// TIA Portal project "Test_PID_Level" (V15.1)

(* hardware
DEVICE "S71500/ET200MP station_1"  S7-1500 station
   slot 0: "Telaio di montaggio_0"  Rack  6ES7 590-1***0-0AA0
   slot 1: "PLC_1"  CPU 1515-2 PN  6ES7 515-2AM01-0AB0  V2.6
      slot 3: "Display CPU_1"  6ES7591-1BA00-0AA0
DEVICE "HMI_1"  TP2200 Comfort
   slot 0: "HMI_1"  TP2200 Comfort  6AV2 124-0XC02-0AX1  15.1.0.0
   slot 1: "HMI_RT_1"  TP2200 Comfort  6AV2 124-0XC02-0AX1  15.1.0.0
   slot 5: "HMI_1.IE_CP_1"  PROFINET Interface  15.0.1.0
      slot 1: "Interfaccia_1 PROFINET"  PROFINET Interface
         slot 1: "Porta_1"  Port
         slot 2: "Porta_2"  Port
   slot 6: "HMI_1.IE_CP_2"  PROFINET Interface  15.0.1.0
      slot 1: "PROFINET Interface_GBit"  PROFINET Interface
         slot 1: "Porta_1"  Port
   slot 7: "HMI_1.MPI/DP_CP_1"  MPI/DP Interface  15.0.1.0
*)

// ===== PLC "PLC_1"  CPU 1515-2 PN =====

TYPE "s_PID"
   STRUCT
      i_Set_Point : Real;   // Set point value
      i_Feedback : Real;   // Feedback value process
      i_Kp : Real;   // K Proportional gain
      i_Ki : Real;   // K Integral gain
      i_Kd : Real;   // K Derivative gain
      i_Max_Analog : Real;   // Maximum value for analog output
      i_Duty_Cycle : Real;   // Maximum time cycle for PWM digital output (milliseconds)
      i_Scan_Time : Real;   // Scanning time of the plc
      i_Time_Sample : Real;   // Time sample in OB35
      i_Enable_PWM : Bool;   // Enable PWM digital P.I.D.
      i_Reset : Bool;   // Reset regulator
      i_Enable_I : Bool;   // Enable Integral component
      o_Analog_Reg : Real;   // Output analog regulation
      o_Duty_Cycle_Perc : Real;   // Duty cycle On percentage
      o_Wave_On_PWM : Bool;   // Output high wave On of digital PWM
      o_Wave_Off_PWM : Bool;   // Output low wave On of digital PWM
   END_STRUCT;
END_TYPE

DATA_BLOCK "f_PID_DB"   // DB80
{ S7_Optimized_Access := 'TRUE' }
VERSION : 0.1
// stored: InstanceOfName f_PID
"f_PID"
BEGIN
END_DATA_BLOCK

DATA_BLOCK "DB_PID"   // DB82
{ S7_Optimized_Access := 'TRUE' }
VERSION : 0.1
   VAR RETAIN
      Data : "s_PID";   // Valve 1
   END_VAR
   VAR
      Scan_Time_LR : LReal;
      Mem_Scan_Time : LReal;
      Scan_Time_R : Real;
      FB_Int : Int;
      Derivative_ON : Bool;
      Enable_I : Bool;
   END_VAR
BEGIN
END_DATA_BLOCK

DATA_BLOCK "DB_Tank"   // DB83
{ S7_Optimized_Access := 'TRUE' }
VERSION : 0.1
   VAR
      V1_On : Bool;
      V2_On : Bool;
      V3_On : Bool;
      V4_On : Bool;
      V1_Max : Real;   // Liters per second V1, input
      V2_SP : Real;   // Set point Liters per second
      V3_SP : Real;   // Set point Liters per second
      V4_SP : Real;   // Set point Liters per second
      Water : Real;   // Liters
      Tank_Max : Real := 3000.0;
      V1_In : Real;   // Liters in input
      V2_Out : Real;   // Liters in output
      V3_Out : Real;   // Liters in output
      V4_Out : Real;   // Liters in output
      FB_V1 : Real;
   END_VAR
BEGIN
END_DATA_BLOCK

FUNCTION_BLOCK "f_PID"   // FB80, SCL
{ S7_Optimized_Access := 'TRUE' }
VERSION : 0.1
   VAR_INPUT
      Set_Point : Real;   // Set point value
      Feedback : Real;   // Feedback value process
      Kp : Real;   // K Proportional gain
      Ki : Real;   // K Integral gain
      Kd : Real;   // K Derivative gain
      Max_Analog : Real;   // Maximum value for analog output
      Duty_Cycle : Real;   // Maximum time cycle for PWM digital output (milliseconds)
      Scan_Time : Real;   // Scanning time of the plc
      Time_Sample : Real;   // Time sample in OB35
      Enable_PWM : Bool;   // Enable PWM digital P.I.D.
      Reset : Bool;   // Reset regulator
      Enable_I : Bool;
   END_VAR
   VAR_OUTPUT
      Analog_Reg : Real;   // Output analog regulation
      Duty_Cycle_Perc : Real;   // Duty cycle On percentage
      Wave_On_PWM : Bool;   // Output high wave On of digital PWM
      Wave_Off_PWM : Bool;   // Output low wave On of digital PWM
      Derivative_ON : Bool;
   END_VAR
   VAR
      Error : Real;   // Error for each scan
      I_Ist : Real;   // Istant integral
      I : Real;   // Integral component
      D : Real;   // Derivative component
      P : Real;   // Proportional component
      Last_Error : Real;   // Error of previous scan
      Accu_Timer : Real;   // Timer Accumulator for the duty cycle PWM
      Thr_Wave_On : Real;   // Threshold for the wave ON
      Thr_Wave_Off : Real;   // Threshold for the wave OFF
      Wave_On : Bool;   // Wave On
      Wave_Off : Bool;   // Wave Off
   END_VAR
BEGIN
   // P.I.D. Regulator. Written By Ing. Walter Porcellini Milan (Italy) the 15/09/2021
   // I revisited and modified the algorithm I wrote in June 2009
   // This project and its algorithm are intended as a didactic demonstration
   // I decline from any responsibility for damage to things and / or people.

   #Error := #Set_Point - #Feedback;

   #P := #Error * #Kp * 1.0;

   IF #P > #Max_Analog THEN

       #P := #Max_Analog;
   END_IF;

   IF #P < (#Max_Analog * -1.0) THEN

       #P := #Max_Analog * -1.0;
   END_IF;

   IF #Enable_I = true THEN
       #I_Ist := #Error * #Ki * 1.0;
       #I := #I + #I_Ist;

   ELSE
       #I_Ist := 0.0;
       #I := 0.0;
   END_IF;

   #I := #I + #I_Ist;

   IF #I <= 0.0 THEN
      #I := 0.0;
   END_IF;

   IF #I >= #Max_Analog * 0.8 THEN
       #I := #Max_Analog * 0.8;
   END_IF;

   IF #Time_Sample > 0.0 THEN
       #D := (#Kd * 1.0*(#Error - #Last_Error)) / #Time_Sample;
   END_IF;

   #Last_Error := #Error;

   #Analog_Reg := #P + #I + #D;

   #Derivative_ON := #D <> 0.0;

   IF #Reset THEN

       #P := 0.0;
       #I := 0.0;
       #I_Ist := 0.0;
       #D := 0.0;
       #Analog_Reg := 0.0;
       #Wave_On := false;
       #Wave_Off := false;
       #Accu_Timer := 0.0;
       #Last_Error := 0.0;

   END_IF;

   IF #Analog_Reg >= #Max_Analog THEN
       #Analog_Reg := #Max_Analog;
   END_IF;

   IF #Analog_Reg <= 0.0 THEN
       #Analog_Reg:=0.0;
   END_IF;


   IF #Enable_PWM = true THEN
       #Thr_Wave_On := (#Duty_Cycle / #Max_Analog) * #Analog_Reg;

       #Thr_Wave_Off := #Max_Analog - #Thr_Wave_On;


       IF #Accu_Timer = 0.0 AND #Enable_PWM = TRUE THEN

           #Wave_On := true;
           #Wave_Off := false;

       END_IF;

       IF #Wave_On = true THEN

           #Accu_Timer := #Accu_Timer + #Time_Sample;
           #Duty_Cycle_Perc := (#Thr_Wave_On / #Duty_Cycle) * 100.0;

           IF #Accu_Timer >= #Thr_Wave_On THEN

               #Wave_On := false;
               #Wave_Off := true;

           END_IF;

       END_IF;


       IF #Wave_Off = true THEN

           #Accu_Timer := #Accu_Timer + #Time_Sample;

           IF #Accu_Timer >= #Duty_Cycle THEN

               #Wave_Off := false;
               #Accu_Timer := 0.0;

           END_IF;

       END_IF;



       #Wave_On_PWM := #Wave_On AND #Thr_Wave_On >= 1000.0;
       #Wave_Off_PWM := #Wave_Off;

   ELSE
       #Wave_On_PWM := false;
       #Wave_Off_PWM := false;
       #Accu_Timer := 0.0;
       #Duty_Cycle_Perc := 0.0;
   END_IF;
END_FUNCTION_BLOCK

FUNCTION "1_Temperature" : Void   // FC100, SCL
{ S7_Optimized_Access := 'TRUE' }
VERSION : 0.1
BEGIN
   // "DB_PID".V1.i_Feedback := INT_TO_REAL("DB_PID".FB_Int);

   "DB_PID".Data.i_Feedback := "DB_PID".Data.i_Feedback + ("DB_PID".Data.o_Analog_Reg * 0.000000024);
   "DB_PID".Data.i_Feedback := "DB_PID".Data.i_Feedback - 0.00008;

   IF "DB_PID".Data.i_Feedback < 20.0 OR "DB_PID".Data.i_Reset = true THEN

       "DB_PID".Data.i_Feedback := 20.0;
   END_IF;


   IF "DB_PID".Data.i_Feedback > 150.0 THEN

       "DB_PID".Data.i_Feedback := 150.0;
   END_IF;
END_FUNCTION

FUNCTION "2_Tank Level" : Void   // FC101, SCL
{ S7_Optimized_Access := 'TRUE' }
VERSION : 0.1
   VAR_TEMP
      Stop_Integral : Bool;
   END_VAR
BEGIN

   IF "DB_Tank".V2_SP > 30.0 THEN

       "DB_Tank".V2_SP := 30.0;

   END_IF;

   IF "DB_Tank".V2_SP < 0.0 THEN

       "DB_Tank".V2_SP := 0.0;

   END_IF;

   IF "DB_Tank".V3_SP > 30.0 THEN

       "DB_Tank".V3_SP := 30.0;

   END_IF;

   IF "DB_Tank".V3_SP < 0.0 THEN

       "DB_Tank".V3_SP := 0.0;

   END_IF;

   IF "DB_Tank".V4_SP > 30.0 THEN

       "DB_Tank".V4_SP := 30.0;

   END_IF;

   IF "DB_Tank".V4_SP < 0.0 THEN

       "DB_Tank".V4_SP := 0.0;

   END_IF;

   "DB_Tank".V2_Out := ("DB_Tank".V2_SP * "DB_PID".Scan_Time_R);
   "DB_Tank".V3_Out := ("DB_Tank".V3_SP * "DB_PID".Scan_Time_R);
   "DB_Tank".V4_Out := ("DB_Tank".V4_SP * "DB_PID".Scan_Time_R);

   IF "DB_Tank".V2_On = true THEN
       "DB_Tank".Water := "DB_Tank".Water - "DB_Tank".V2_Out;

   END_IF;

   IF "DB_Tank".V3_On = true THEN
       "DB_Tank".Water := "DB_Tank".Water - "DB_Tank".V3_Out;

   END_IF;

   IF "DB_Tank".V4_On = true THEN
       "DB_Tank".Water := "DB_Tank".Water - "DB_Tank".V4_Out;

   END_IF;

   "DB_Tank".V1_Max := 100.0;
   "DB_Tank".V1_In := ("DB_Tank".V1_Max / "DB_PID".Data.i_Max_Analog) * "DB_PID".Data.o_Analog_Reg * "DB_PID".Scan_Time_R ;
   "DB_Tank".FB_V1 := "DB_Tank".V1_In * 1000.0;

   "DB_Tank".Water := "DB_Tank".Water + "DB_Tank".V1_In;

   IF "DB_Tank".Water < 0.0 OR "DB_PID".Data.i_Reset=true THEN

       "DB_Tank".Water := 0;
   END_IF;

   "DB_Tank".V1_On := "DB_PID".Data.o_Analog_Reg > 0.0;
   "DB_PID".Data.i_Feedback := "DB_Tank".Water;
   "DB_PID".FB_Int := REAL_TO_INT("DB_Tank".Water);

   #Stop_Integral := "DB_Tank".V2_On = false
   AND "DB_Tank".V3_On = false
   AND "DB_Tank".V4_On = false;

   "DB_PID".Enable_I := NOT #Stop_Integral;
END_FUNCTION

ORGANIZATION_BLOCK "Main"   // OB1, LAD, ProgramCycle
TITLE = "Main Program Sweep (Cycle)"
{ S7_Optimized_Access := 'TRUE' }
VERSION : 0.1
   VAR_INPUT
      Initial_Call : Bool;   // Initial call of this OB
      Remanence : Bool;   // =True, if remanent data are available
   END_VAR
BEGIN

REGION Network 1
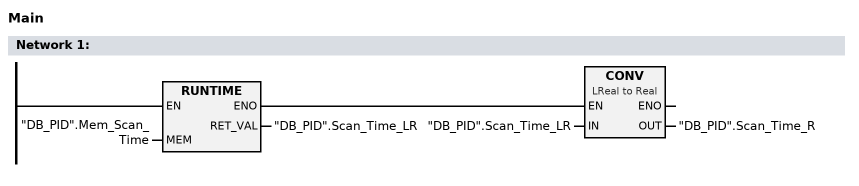
   // no SCL statement known for Runtime: written as a call
   // ENO of a box is taken as its EN; it also drops when the box reports an error
   "DB_PID".Scan_Time_LR := Runtime(mem := "DB_PID".Mem_Scan_Time);
   "DB_PID".Scan_Time_R := LREAL_TO_REAL("DB_PID".Scan_Time_LR);
END_REGION

REGION Network 2 (SCL)
   "DB_PID".Data.i_Max_Analog := 16384;
   "DB_PID".Data.i_Duty_Cycle := 10000;
   "DB_PID".Data.i_Scan_Time := "DB_PID".Scan_Time_R;
   "DB_PID".Data.i_Time_Sample := 10;

   //"1_Temperature"();
   "2_Tank Level"();
END_REGION
END_ORGANIZATION_BLOCK

ORGANIZATION_BLOCK "Cyclic interrupt"   // OB30, LAD, CyclicInterrupt
{ S7_Optimized_Access := 'TRUE' }
VERSION : 0.1
   VAR_INPUT
      Initial_Call : Bool;   // Initial call of this OB
      Event_Count : Int;   // Events discarded
   END_VAR
BEGIN

REGION Network 1
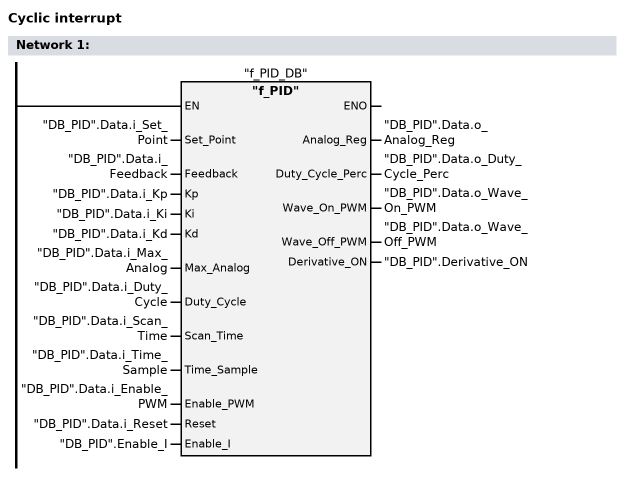
   RUNG wire#powerrail
      "f_PID_DB"(Set_Point := "DB_PID".Data.i_Set_Point, Feedback := "DB_PID".Data.i_Feedback, Kp := "DB_PID".Data.i_Kp, Ki := "DB_PID".Data.i_Ki, Kd := "DB_PID".Data.i_Kd, Max_Analog := "DB_PID".Data.i_Max_Analog, Duty_Cycle := "DB_PID".Data.i_Duty_Cycle, Scan_Time := "DB_PID".Data.i_Scan_Time, Time_Sample := "DB_PID".Data.i_Time_Sample, Enable_PWM := "DB_PID".Data.i_Enable_PWM, Reset := "DB_PID".Data.i_Reset, Enable_I := "DB_PID".Enable_I, Analog_Reg => "DB_PID".Data.o_Analog_Reg, Duty_Cycle_Perc => "DB_PID".Data.o_Duty_Cycle_Perc, Wave_On_PWM => "DB_PID".Data.o_Wave_On_PWM, Wave_Off_PWM => "DB_PID".Data.o_Wave_Off_PWM, Derivative_ON => "DB_PID".Derivative_ON)
   END_RUNG
   // the same network as SCL:
   "f_PID_DB"(Set_Point := "DB_PID".Data.i_Set_Point,   // "f_PID"
              Feedback := "DB_PID".Data.i_Feedback,
              Kp := "DB_PID".Data.i_Kp,
              Ki := "DB_PID".Data.i_Ki,
              Kd := "DB_PID".Data.i_Kd,
              Max_Analog := "DB_PID".Data.i_Max_Analog,
              Duty_Cycle := "DB_PID".Data.i_Duty_Cycle,
              Scan_Time := "DB_PID".Data.i_Scan_Time,
              Time_Sample := "DB_PID".Data.i_Time_Sample,
              Enable_PWM := "DB_PID".Data.i_Enable_PWM,
              Reset := "DB_PID".Data.i_Reset,
              Enable_I := "DB_PID".Enable_I,
              Analog_Reg => "DB_PID".Data.o_Analog_Reg,
              Duty_Cycle_Perc => "DB_PID".Data.o_Duty_Cycle_Perc,
              Wave_On_PWM => "DB_PID".Data.o_Wave_On_PWM,
              Wave_Off_PWM => "DB_PID".Data.o_Wave_Off_PWM,
              Derivative_ON => "DB_PID".Derivative_ON);
END_REGION
END_ORGANIZATION_BLOCK

(* ===== HMI "HMI_RT_1" =====
system functions are stored by id; their names below are inferred from use
connection "HMI_Collegamento_1": ETHERNET, S7_1500_OMS

HMI tags "Tabella delle variabili standard"
   "Variabile_Numero di pagina" : UInt, internal
   "DB_PID_V1_i_Set_Point" : Real = PLC DB_PID.Data.i_Set_Point, 1 s
   "DB_PID_V1_i_Kp" : Real = PLC DB_PID.Data.i_Kp, 1 s
   "DB_PID_V1_i_Feedback" : Real = PLC DB_PID.Data.i_Feedback, 1 s
   "DB_PID_V1_i_Ki" : Real = PLC DB_PID.Data.i_Ki, 1 s
   "DB_PID_V1_i_Kd" : Real = PLC DB_PID.Data.i_Kd, 1 s
   "DB_PID_V1_i_Enable_PWM" : Bool = PLC DB_PID.Data.i_Enable_PWM, 1 s
   "DB_PID_V1_i_Reset" : Bool = PLC DB_PID.Data.i_Reset, 1 s
   "DB_PID_V1_o_Analog_Reg" : Real = PLC DB_PID.Data.o_Analog_Reg, 1 s
   "DB_PID_V1_o_Duty_Cycle_Perc" : Real = PLC DB_PID.Data.o_Duty_Cycle_Perc, 1 s
   "DB_PID_V1_o_Wave_On_PWM" : Bool = PLC DB_PID.Data.o_Wave_On_PWM, 1 s
   "DB_PID_V1_o_Wave_Off_PWM" : Bool = PLC DB_PID.Data.o_Wave_Off_PWM, 1 s
   "DB_PID_FB_Int" : Int = PLC DB_PID.FB_Int, 1 s
   "DB_PID_Derivative_ON" : Bool = PLC DB_PID.Derivative_ON, 1 s
   "DB_Tank_V1_On" : Bool = PLC DB_Tank.V1_On, 1 s
   "DB_Tank_V2_On" : Bool = PLC DB_Tank.V2_On, 1 s
   "DB_Tank_V3_On" : Bool = PLC DB_Tank.V3_On, 1 s
   "DB_Tank_V4_On" : Bool = PLC DB_Tank.V4_On, 1 s
   "DB_Tank_V2_SP" : Real = PLC DB_Tank.V2_SP, 1 s
   "DB_Tank_V3_SP" : Real = PLC DB_Tank.V3_SP, 1 s
   "DB_Tank_V4_SP" : Real = PLC DB_Tank.V4_SP, 1 s
   "f_PID_DB_P" : Real = PLC f_PID_DB.P, 1 s
   "f_PID_DB_I" : Real = PLC f_PID_DB.I, 1 s
   "f_PID_DB_D" : Real = PLC f_PID_DB.D, 1 s
   "DB_Tank_V1_In" : Real = PLC DB_Tank.V1_In, 1 s
   "DB_Tank_FB_V1" : Real = PLC DB_Tank.FB_V1, 1 s

text list "Elenco testi_Nome della pagina": 1 'Pagina base'

screen "Pagina base" 1920x1017, template "Modello_1"
   on GenerateScreen: SetTag("Variabile_Numero di pagina", 1)
   TextField "Casella di testo_1" at 9,24 size 98x25; Text 'Set Point'
   IOField "Campo I/O_1" at 114,21 size 96x32; FormatPattern 9999.9
      ProcessValue <- "DB_PID_V1_i_Set_Point"
   TextField "Casella di testo_2" at 9,68 size 30x25; Text 'Kp'
   IOField "Campo I/O_2" at 114,64 size 96x32; FormatPattern 9999.9
      ProcessValue <- "DB_PID_V1_i_Kp"
   TextField "Casella di testo_3" at 9,111 size 24x25; Text 'Ki'
   IOField "Campo I/O_3" at 114,108 size 96x32; FormatPattern 9999.9
      ProcessValue <- "DB_PID_V1_i_Ki"
   TextField "Casella di testo_4" at 9,155 size 30x25; Text 'Kd'
   IOField "Campo I/O_4" at 114,151 size 96x32; FormatPattern 9999.9
      ProcessValue <- "DB_PID_V1_i_Kd"
   TextField "Casella di testo_8" at 354,24 size 94x25; Text 'Feedback'
   IOField "Campo I/O_5" at 255,21 size 96x32; FormatPattern 9999.9
      ProcessValue <- "DB_PID_V1_i_Feedback"
   Switch "Interruttore_1" at 100,197 size 120x67; CaptionText 'Enable PWM'; TextOff 'OFF'; TextOn 'ON'
      ProcessValue <- "DB_PID_V1_i_Enable_PWM"
   Switch "Interruttore_2" at 100,269 size 120x67; TextOn 'ON'; CaptionText 'Reset'; TextOff 'OFF'
      ProcessValue <- "DB_PID_V1_i_Reset"
   TextField "Casella di testo_5" at 579,66 size 143x25; Text 'Analog Output'
   IOField "Campo I/O_6" at 475,64 size 96x32; FormatPattern s99999
      ProcessValue <- "DB_PID_V1_o_Analog_Reg"
   TextField "Casella di testo_6" at 579,217 size 77x25; Text 'Duty %'
   IOField "Campo I/O_7" at 475,215 size 96x32; FormatPattern 9999.9
      ProcessValue <- "DB_PID_V1_o_Duty_Cycle_Perc"
   Ellipse "Ellisse_1" at 538,258 size 30x30
      Appearance <- "DB_PID_V1_o_Wave_On_PWM"
   TextField "Casella di testo_9" at 579,262 size 85x25; Text 'PWM ON'
   Bar "Barra grafica_1" at 475,21 size 151x36; MinimumValue 0; MaximumValue 16384
      ProcessValue <- "DB_PID_V1_o_Analog_Reg"
   GraphicView "Vista grafica_2" at 1028,62 size 300x260; Picture "Grafica_2"
   Bar "Barra grafica_2" at 1051,141 size 249x174; MinimumValue 0; MaximumValue 3000
      ProcessValue <- "DB_PID_FB_Int"
   GraphicView "Vista grafica_3" at 892,19 size 96x43; Picture "valvola_off_1"
   GraphicView "Vista grafica_1" at 893,19 size 96x43; Picture "valvola_on"
      Visibility <- "DB_Tank_V1_On"
   GraphicView "Vista grafica_4" at 893,264 size 96x43; Picture "valvola_off_1"
   GraphicView "Vista grafica_5" at 893,264 size 96x43; Picture "valvola_on"
      Visibility <- "DB_Tank_V2_On"
   GraphicView "Vista grafica_10" at 1356,270 size 96x43; Picture "valvola_off_1"
   GraphicView "Vista grafica_11" at 1356,270 size 96x43; Picture "valvola_on"
      Visibility <- "DB_Tank_V3_On"
   GraphicView "Vista grafica_12" at 1186,378 size 96x43; Picture "valvola_off_1"
   GraphicView "Vista grafica_13" at 1186,378 size 96x43; Picture "valvola_on"
      Visibility <- "DB_Tank_V4_On"
   Button "Pulsante_1" at 1462,194 size 96x32; TextOff 'ON'
      on Press: SetBit("DB_Tank_V3_On")
   Button "Pulsante_2" at 1463,227 size 96x32; TextOff 'OFF'
      on Press: ResetBit("DB_Tank_V3_On")
   Button "Pulsante_3" at 893,338 size 96x32; TextOff 'ON'
      on Press: SetBit("DB_Tank_V2_On")
   Button "Pulsante_4" at 894,371 size 96x32; TextOff 'OFF'
      on Press: ResetBit("DB_Tank_V2_On")
   Button "Pulsante_5" at 1355,366 size 96x32; TextOff 'ON'
      on Press: SetBit("DB_Tank_V4_On")
   Button "Pulsante_6" at 1356,399 size 96x32; TextOff 'OFF'
      on Press: ResetBit("DB_Tank_V4_On")
   IOField "Campo I/O_8" at 892,68 size 96x32; FormatPattern 9999.9
      ProcessValue <- "DB_Tank_FB_V1"
   IOField "Campo I/O_9" at 893,229 size 96x32; FormatPattern 9999.9
      ProcessValue <- "DB_Tank_V2_SP"
   IOField "Campo I/O_10" at 1356,231 size 96x32; FormatPattern 9999.9
      ProcessValue <- "DB_Tank_V3_SP"
   IOField "Campo I/O_11" at 1186,346 size 96x32; FormatPattern 9999.9
      ProcessValue <- "DB_Tank_V4_SP"
   GraphicView "Vista grafica_6" at 1497,284 size 41x21; Picture "Right_Arrow"
   GraphicView "Vista grafica_7" at 804,275 size 41x21; Picture "Left_Arrow"
   GraphicView "Vista grafica_14" at 809,30 size 41x21; Picture "Right_Arrow"
   GraphicView "Vista grafica_15" at 1282,388 size 41x21; Picture "Right_Arrow"
   TextField "Casella di testo_7" at 362,68 size 17x25; Text 'P'
   IOField "Campo I/O_12" at 255,64 size 96x32; FormatPattern 999999
      ProcessValue <- "f_PID_DB_P"
   TextField "Casella di testo_10" at 362,111 size 14x25; Text 'I'
   IOField "Campo I/O_13" at 255,108 size 96x32; FormatPattern 999999
      ProcessValue <- "f_PID_DB_I"
   IOField "Campo I/O_14" at 255,151 size 96x32; FormatPattern s99999
      ProcessValue <- "f_PID_DB_D"
   TextField "Casella di testo_11" at 362,155 size 19x25; Text 'D'
   TextField "Casella di testo_12" at 627,26 size 91x25; Text '(0 -10 V)'
   TextField "Casella di testo_13" at 1366,203 size 72x25; Text 'L / Sec'
   TextField "Casella di testo_14" at 905,102 size 72x25; Text 'L / Sec'
   TextField "Casella di testo_15" at 905,203 size 72x25; Text 'L / Sec'
   TextField "Casella di testo_16" at 1199,318 size 72x25; Text 'L / Sec'

Template "Modello_1" 1920x1017
   Button "Esci" at 720,360 size 78x58; TextOff 'Esci'; PictureOff "ExitRuntime_TP900_Comfort_TR"; PictureOn "ExitRuntime_TP900_Comfort_TR"
      on Release: StopRuntime(0)
   Button "Template_Button" at 640,360 size 78x58; TextOff 'Text'
   Button "Template_Button_1" at 560,360 size 78x58; TextOff 'Text'
   Button "Template_Button_2" at 480,360 size 78x58; TextOff 'Text'
   Button "Template_Button_3" at 400,360 size 78x58; TextOff 'Text'
   Button "Template_Button_4" at 321,360 size 78x58; TextOff 'Text'
   Button "Template_Button_5" at 241,360 size 78x58; TextOff 'Text'
   Button "Template_Button_6" at 161,360 size 78x58; TextOff 'Text'
   Button "Segnalazioni" at 81,360 size 78x58; TextOff 'Segnalazioni'; PictureOff "AlarmDisplay_TP900_Comfort_TR"; PictureOn "AlarmDisplay_TP900_Comfort_TR"
      on Release: function_ef3f5d25("Finestra delle segnalazioni_Non riconosciuta", -1)
   Button "Pagina iniziale" at 1,360 size 78x58; TextOff 'Pagina iniziale'; PictureOff "NavigateHome_TP900_Comfort_TR"; PictureOn "NavigateHome_TP900_Comfort_TR"
      on Release: ActivateScreen("Pagina base", 0)
*)